      Visibility <- "10_DI_DATA_FS_332 FLW_OK"
      HorizontalMovement <- "82_To_HMI_FS332 Animation"
   Circle "Circle_69" at 573,764 size 8x8
      Visibility <- "10_DI_DATA_FS_332 FLW_OK"
      HorizontalMovement <- "82_To_HMI_FS332 Animation"
   Circle "Circle_70" at 712,763 size 8x8
      Visibility <- "10_DI_DATA_FS_332 FLW_OK"
      HorizontalMovement <- "82_To_HMI_FS332 Animation"
   Circle "Circle_74" at 822,763 size 8x8
      Visibility <- "10_DI_DATA_FS_332 FLW_OK"
      HorizontalMovement <- "82_To_HMI_FS332 Animation"
   Circle "Circle_75" at 828,691 size 8x8
      Visibility <- "10_DI_DATA_FS_332 FLW_OK"
      VerticalMovement <- "82_To_HMI_FS332 Animation"
   Circle "Circle_76" at 828,633 size 8x8
      Visibility <- "10_DI_DATA_FS_332 FLW_OK"
      VerticalMovement <- "82_To_HMI_FS332 Animation"
   Circle "Circle_77" at 763,613 size 8x8
      Visibility <- "10_DI_DATA_FS_332 FLW_OK"
      HorizontalMovement <- "82_To_HMI_FS332 Animation"
   Circle "Circle_78" at 845,515 size 10x10
      Visibility <- "10_DI_DATA_FS_332 FLW_OK"
      HorizontalMovement <- "82_To_HMI_FS332 Animation"
   Circle "Circle_79" at 856,642 size 10x10
      Visibility <- "10_DI_DATA_FS_332 FLW_OK"
      VerticalMovement <- "82_To_HMI_FS332 Animation"
   Circle "Circle_80" at 856,765 size 10x10
      Visibility <- "10_DI_DATA_FS_332 FLW_OK"
      VerticalMovement <- "82_To_HMI_FS332 Animation"
   Circle "Circle_55" at 179,684 size 7x7
      Visibility <- "10_DI_DATA_CV358_OPN"
      HorizontalMovement <- "82_To_HMI_P304 Animation"
   Circle "Circle_83" at 318,685 size 7x7
      Visibility <- "10_DI_DATA_CV358_OPN"
      DiagonalMovement <- "82_To_HMI_P304 Animation"
   Circle "Circle_81" at 416,684 size 7x7
      Visibility <- "10_DI_DATA_CV358_OPN"
      DiagonalMovement <- "82_To_HMI_P304 Animation"
   Circle "Circle_56" at 485,684 size 7x7
      Visibility <- "10_DI_DATA_CV358_OPN"
      DiagonalMovement <- "82_To_HMI_P304 Animation"
   Circle "Circle_85" at 496,641 size 7x7
      Visibility <- "10_DI_DATA_CV358_OPN"
      DiagonalMovement <- "82_To_HMI_P304 Animation"
   Circle "Circle_86" at 426,634 size 7x7
      Visibility <- "10_DI_DATA_CV358_OPN"
      DiagonalMovement <- "82_To_HMI_P304 Animation"
   TextField "Text field_50" at 969,420 size 254x154; Text 'Please Make Sure the Energy and Water Supply are Present and Sufficient'
      Visibility <- "Warn To Start GCU-Last"
   Button "Button_5" at 928,406 size 343x378; TextOff 'Text'
      Visibility <- "Warn To Start GCU-Last"
   TextField "Text field_21" at 919,606 size 359x94; Text 'Instalation Start Confirmation Required for Re-Ox Stage'
      Visibility <- "Warn To Start GCU-Last"
   Button "Button_6" at 1004,717 size 200x55; TextOff 'CONFIRM'; Authorization "Operate"
      on Press: function_b14e0dd5("80_From_HMI_GCU Start Confirmed", 0)
      Visibility <- "Warn To Start GCU-Last"
   TextField "Text field_51" at 914,433 size 366x124; Text 'Please Make Sure the Energy and Water Supply are Present and Sufficient'
      Visibility <- "Warn To Start GCU-Last"
   IOField "I/O field_37" at 1070,718 size 79x29; Authorization "Commissioning"; FormatPattern 999; Unit  step
      ProcessValue <- "2110_BTCS_CNTRL_DB_BTCS_STEP"
   Button "HmiScreenItemData_18" at 930,718 size 137x29; TextOn 'Back'; TextOff 'BWTS Step'
   Button "HmiScreenItemData_51" at 930,753 size 137x29; TextOn 'Back'; TextOff 'BWTS State'
   IOField "I/O field_38" at 1070,753 size 79x29; Authorization "Commissioning"; FormatPattern 9; Unit  state
      ProcessValue <- "2110_BTCS_CNTRL_DB_BTCS_STATE"
   TextField "Text field_64" at 497,462 size 54x22; Text '- OK -'
      Visibility <- "10_DI_DATA_LS_303_LO"
   GraphicView "Graphic view_76" at 53,433 size 168x182; Picture "Graphic_251"
   GraphicView "Graphic view_102" at 12,304 size 58x63; Picture "Graphic_162"
   GraphicView "Graphic view_13" at 724,163 size 182x22; Picture "Graphic_151"
   GraphicIOField "Graphic I/O field_3" at 188,659 size 60x65; PictureList "Pump Ani"
      ProcessValue <- "10_DI_DATA_P_304_ENBLD"
   GraphicView "Graphic view_18" at 240,683 size 253x11; Picture "Graphic_156"
   GraphicView "Graphic view_89" at 303,257 size 10x13; Picture "Graphic_147"
   GraphicView "Graphic view_59" at 962,301 size 302x22; Picture "Graphic_151"
   GraphicView "Graphic view_5" at 827,163 size 102x22; Picture "Graphic_151"
   GraphicView "Graphic view_69" at 124,683 size 68x11; Picture "Graphic_156"
   GraphicView "Graphic view_85" at 235,296 size 33x35; Picture "Graphic_178"
   GraphicView "Graphic view_1" at 259,128 size 301x502; Picture "Graphic_150"
   GraphicView "Graphic view_6" at 870,257 size 18x22; Picture "Graphic_154"
   GraphicView "Graphic view_9" at 689,257 size 188x11; Picture "Graphic_156"
   GraphicView "Graphic view_11" at 424,625 size 12x91; Picture "Graphic_152"
   GraphicView "Graphic view_10" at 424,628 size 19x28; Picture "Graphic_157"
   GraphicView "Graphic view_12" at 440,636 size 106x11; Picture "Graphic_156"
   GraphicView "Graphic view_14" at 817,752 size 20x21; Picture "Graphic_159"
   GraphicView "Graphic view_16" at 635,761 size 188x13; Picture "Graphic_151"
   GraphicIOField "Graphic I/O field_1" at 573,615 size 60x65; PictureList "Pump Ani"
      ProcessValue <- "10_DI_DATA_P_303_ENBLD"
   GraphicView "Graphic view_19" at 471,636 size 106x11; Picture "Graphic_156"
   TextField "Text field_16" at 90,573 size 90x22; Text 'PGC Running'
      Visibility <- "10_DI_DATA_E_400_RUN"
   GraphicView "Graphic view_21" at 486,674 size 17x18; Picture "Graphic_153"
   GraphicView "Graphic view_22" at 494,642 size 10x41; Picture "Graphic_152"
   GraphicView "Graphic view_23" at 490,637 size 17x15; Picture "Graphic_161"
   GraphicView "Graphic view_24" at 630,636 size 87x11; Picture "Graphic_156"
   GraphicView "Graphic view_33" at 668,469 size 24x18; Picture "Graphic_155"
   GraphicView "Graphic view_34" at 668,508 size 24x18; Picture "Graphic_166"
   GraphicView "Graphic view_35" at 679,517 size 62x11; Picture "Graphic_156"
   GraphicView "Graphic view_36" at 668,486 size 12x30; Picture "Graphic_152"
   GraphicView "Graphic view_37" at 687,468 size 62x11; Picture "Graphic_156"
   GraphicView "Graphic view_38" at 741,468 size 106x11; Picture "Graphic_156"
   GraphicView "Graphic view_39" at 487,257 size 103x11; Picture "Graphic_156"
   GraphicView "Graphic view_40" at 422,102 size 140x11; Picture "Graphic_156"
   GraphicView "Graphic view_41" at 302,103 size 24x18; Picture "Graphic_155"
   GraphicView "Graphic view_43" at 558,103 size 19x18; Picture "Graphic_154"
   GraphicView "Graphic view_44" at 302,118 size 12x75; Picture "Graphic_152"
   GraphicView "Graphic view_45" at 302,183 size 12x75; Picture "Graphic_152"
   GraphicView "Graphic view_46" at 871,460 size 17x18; Picture "Graphic_153"
   GraphicView "Graphic view_47" at 879,426 size 10x41; Picture "Graphic_152"
   GraphicView "Graphic view_48" at 771,468 size 106x11; Picture "Graphic_156"
   GraphicView "Graphic view_49" at 879,358 size 10x91; Picture "Graphic_152"
   GraphicView "Graphic view_51" at 879,272 size 10x91; Picture "Graphic_152"
   GraphicView "Graphic view_53" at 574,257 size 126x11; Picture "Graphic_156"
   GraphicView "Graphic view_57" at 319,102 size 140x11; Picture "Graphic_156"
   GraphicView "Graphic view_58" at 1062,188 size 19x119; Picture "Graphic_147"
   TextField "Text field_6" at 995,322 size 50x16; Text 'CV-407'
   GraphicView "Graphic view_61" at 561,250 size 23x16; Picture "Graphic_168"
   GraphicView "Graphic view_62" at 567,179 size 10x77; Picture "Graphic_152"
   TextField "Text field_8" at 1103,322 size 50x16; Text 'CV-411'
   TextField "Text field_13" at 1115,180 size 60x22; Text 'Opened'
      Visibility <- "10_DI_DATA_CV409_OPN"
   TextField "Text field_17" at 582,680 size 42x16; Text 'P-303'
   GraphicView "Graphic view_66" at 508,761 size 188x13; Picture "Graphic_151"
   GraphicView "Graphic view_67" at 375,761 size 188x13; Picture "Graphic_151"
   GraphicView "Graphic view_31" at 424,748 size 12x38; Picture "Graphic_152"
   GraphicView "Graphic view_68" at 118,761 size 285x13; Picture "Graphic_151"
   GraphicView "Graphic view_70" at 826,617 size 12x146; Picture "Graphic_147"
   GraphicView "Graphic view_71" at 818,611 size 19x21; Picture "Graphic_169"
   GraphicView "Graphic view_73" at 14,359 size 19x222; Picture "Graphic_147"
   GraphicView "Graphic view_75" at 696,479 size 76x194; Picture "Graphic_173"
   GraphicView "Graphic view_72" at 760,610 size 68x13; Picture "Graphic_151"
   GraphicView "Graphic view_32" at 847,514 size 19x20; Picture "Graphic_169"
   GraphicView "Graphic view_77" at 759,513 size 97x13; Picture "Graphic_151"
   GraphicView "Graphic view_28" at 855,527 size 12x146; Picture "Graphic_147"
   GraphicView "Graphic view_79" at 855,649 size 12x130; Picture "Graphic_147"
   TextField "Text field_24" at 610,79 size 50x16; Text 'CV-405'
   TextField "Text field_27" at 820,266 size 48x16; Text 'FS-350'
   GraphicView "Graphic view_15" at 834,232 size 20x26; Picture "Graphic_79"
   TextField "Text field_40" at 813,209 size 70x22; Text 'No Flow'
      Visibility <- "10_DI_DATA_FS_350_FLW_OK"
   TextField "Text field_41" at 813,209 size 70x22; Text '- Flow -'
      Visibility <- "10_DI_DATA_FS_350_FLW_OK"
   GraphicView "Graphic view_8" at 558,596 size 10x11; Picture "Graphic_159"
   GraphicView "Graphic view_17" at 563,440 size 5x162; Picture "Graphic_147"
   GraphicView "Graphic view_25" at 558,275 size 10x11; Picture "Graphic_169"
   GraphicView "Graphic view_27" at 563,280 size 5x177; Picture "Graphic_147"
   GraphicView "Graphic view_29" at 486,602 size 78x5; Picture "Graphic_151"
   GraphicView "Graphic view_80" at 488,275 size 76x5; Picture "Graphic_151"
   IOField "I/O field_2" at 524,401 size 82x35; FormatPattern 999.9; Unit  %
      ProcessValue <- "12_AI_Data_LIT_304_SCALED"
   TextField "Text field_29" at 669,184 size 56x16; Text 'PIT-416'
   GraphicView "Graphic view_81" at 687,140 size 20x26; Picture "Graphic_36"
   TextField "Text field_25" at 752,442 size 56x16; Text 'TIT-408'
   TextField "Text field_30" at 512,199 size 56x16; Text 'TIT-406'
   GraphicView "Graphic view_82" at 530,137 size 20x26; Picture "Graphic_36"
   TextField "Text field_26" at 824,348 size 56x16; Text 'PIT-353'
   GraphicView "Graphic view_84" at 15,559 size 33x36; Picture "Graphic_177"
   TextField "Text field_7" at 750,184 size 50x16; Text 'CV-406'
   Bar "Bar_1" at 377,282 size 109x327; Unit  %; MinimumValue 0; MaximumValue 100
      ProcessValue <- "12_AI_Data_LIT_304_SCALED"
   TextField "Text field_48" at 16,624 size 112x20; Text 'PG Compressor'
      Appearance <- "10_DI_DATA_E_400_NOK"
   TextField "Text field_34" at 615,534 size 79x34; Text 'Heat Exchanger'
   TextField "Text field_35" at 551,697 size 100x34; Text 'Recirculation Pump'
   TextField "Text field_36" at 402,782 size 61x18; Text 'To Bilge'
   TextField "Text field_37" at 814,782 size 100x18; Text 'To Overboard'
   TextField "Text field_38" at 571,440 size 55x16; Text 'LIT-304'
   TextField "Text field_39" at 269,693 size 56x16; Text 'PIT-358'
   GraphicView "Graphic view_90" at 287,658 size 20x26; Picture "Graphic_36"
   TextField "Text field_28" at 704,774 size 56x16; Text 'PIT-348'
   GraphicView "Graphic view_83" at 722,736 size 20x26; Picture "Graphic_36"
   TextField "Text field_31" at 778,623 size 48x16; Text 'FS-332'
   GraphicView "Graphic view_91" at 801,585 size 20x26; Picture "Graphic_79"
   TextField "Text field_32" at 779,562 size 70x22; Text 'No Flow'
      Visibility <- "10_DI_DATA_FS_332 FLW_OK"
   TextField "Text field_42" at 779,562 size 70x22; Text '- Flow -'
      Visibility <- "10_DI_DATA_FS_332 FLW_OK"
   TextField "Text field_43" at 197,724 size 42x16; Text 'P-304'
   TextField "Text field_44" at 169,740 size 106x20; Text 'Booster Pump'
   GraphicView "Graphic view_2" at 553,163 size 182x22; Picture "Graphic_151"
   GraphicView "Graphic view_7" at 251,453 size 24x21; Picture "Graphic_107"
   TextField "Text field_46" at 225,501 size 86x16; Text 'E-400-PT002'
   TextField "Text field_47" at 132,408 size 86x16; Text 'E-400-TT002'
   GraphicView "Graphic view_87" at 234,321 size 19x128; Picture "Graphic_147"
   GraphicView "Graphic view_86" at 220,442 size 33x36; Picture "Graphic_159"
   IOField "I/O field_10" at 683,53 size 57x22; FormatPattern 999
      ProcessValue <- "12_AI_Data_CV_405_SCALED"
   IOField "I/O field_11" at 226,482 size 68x18; FormatPattern 999.9; Unit  Bar
      ProcessValue <- "12_AI_Data_E_400_PT002_SCALED"
   IOField "I/O field_13" at 663,119 size 68x18; FormatPattern 99.99; Unit  Bar
      ProcessValue <- "12_AI_Data_PIT_416_SCALED"
   IOField "I/O field_14" at 787,330 size 68x18; FormatPattern 99.99; Unit  Bar
      ProcessValue <- "12_AI_Data_PIT_353_SCALED"
   IOField "I/O field_15" at 704,426 size 68x18; FormatPattern 99.99; Unit  °C
      ProcessValue <- "12_AI_Data_TIT_408_SCALED"
   IOField "I/O field_16" at 698,717 size 68x18; FormatPattern 99.99; Unit  Bar
      ProcessValue <- "12_AI_Data_PIT_348_SCALED"
   IOField "I/O field_7" at 263,638 size 68x18; FormatPattern 99.99; Unit  Bar
      ProcessValue <- "12_AI_Data_PIT_358_SCALED"
   TextField "Text field_57" at 1021,112 size 90x32; Text 'Vent To Atmosphere'
   TextField "Text field_58" at 608,3 size 150x18; Text 'Vent To Atmosphere'
   IOField "I/O field_1" at 143,392 size 68x18; FormatPattern 999.9; Unit  °C
      ProcessValue <- "12_AI_Data_E_400_TE002_SCALED"
   GraphicView "Graphic view_93" at 491,492 size 24x21; Picture "Graphic_107"
   TextField "Text field_63" at 515,491 size 48x16; Text 'LS-303'
   TextField "Text field_66" at 497,462 size 54x22; Text 'Low Low'
      Visibility <- "10_DI_DATA_LS_303_LO"
   TextField "Text field_90" at 497,462 size 54x22; Text '-LOW-'
      Visibility <- "10_DI_DATA_LS_303_LO"
   GraphicView "Graphic view_94" at 99,304 size 58x63; Picture "Graphic_162"
   TextField "Text field_70" at 125,264 size 60x22; Text 'Opened'
      Visibility <- "10_DI_DATA_CV441_OPN"
   TextField "Text field_71" at 126,288 size 50x16; Text 'CV-441'
   GraphicView "Graphic view_95" at 103,278 size 19x41; Picture "Graphic_147"
   TextField "Text field_72" at 93,222 size 65x32; Text 'Ambient Air Inlet'
   GraphicView "Graphic view_96" at 86,364 size 36x39; Picture "Graphic_159"
   GraphicView "Graphic view_97" at 28,382 size 70x22; Picture "Graphic_151"
   TextField "Text field_69" at 125,264 size 60x22; Text 'Closed'
      Visibility <- "10_DI_DATA_CV441_CLSD"
   TextField "Text field_12" at 1115,180 size 60x22; Text 'Closed'
      Visibility <- "10_DI_DATA_CV409_CLSD"
   GraphicView "Graphic view_98" at 0,278 size 33x35; Picture "Graphic_169"
   GraphicView "Graphic view_99" at 856,330 size 23x20; Picture "Graphic_255"
   GraphicView "Graphic view_100" at 728,443 size 20x26; Picture "Graphic_36"
   TextField "Text field_18" at 950,356 size 149x23; Text 'Hazardous Area'
   GraphicView "Graphic view_4" at 1204,277 size 20x26; Picture "Graphic_36"
   IOField "I/O field_3" at 1172,257 size 89x18; FormatPattern s99.99; Unit  Bar
      ProcessValue <- "20_TANKS_IP_DATA_RIO_06_FIRST_TANK_DECK_IG_PRESS"
   TextField "Text field_20" at 1186,322 size 56x16; Text 'PIT-415'
   GraphicView "Graphic view_50" at 100,253 size 26x26; Picture "Graphic_261"
   GraphicView "Graphic view_74" at 549,146 size 18x54; Picture "Graphic_281"
   GraphicView "Graphic view_78" at 256,278 size 17x59; Picture "Graphic_281"
   GraphicView "Graphic view_101" at 213,397 size 23x20; Picture "Graphic_255"
   TextField "Text field_56" at 1229,342 size 44x32; Text 'To BWTS'
   TextField "Text field_60" at 661,356 size 94x23; Text 'Safe Area'
   IOField "I/O field_4" at 683,37 size 57x22; FormatPattern 999
      ProcessValue <- "16_AQ_Data_CV405_CNTRL"
   TextField "Text field_106" at 752,38 size 59x18; Text 'OPENED'
   GraphicView "Graphic view_103" at 14,298 size 19x22; Picture "Graphic_147"
   TextField "Text field_73" at 34,288 size 50x16; Text 'CV-401'
   TextField "Text field_74" at 30,264 size 60x22; Text 'Opened'
      Visibility <- "10_DI_Data_CV401_OPN"
   TextField "Text field_75" at 30,264 size 60x22; Text 'Closed'
      Visibility <- "10_DI_Data_CV401_CLSD"
   Button "HmiScreenItemData_13" at 4,669 size 121x40; TextOn 'IGG Plant'; TextOff 'Fresh Water System'
      on Release: ActivateScreen("Fresh Water System", 0)
      Appearance <- "10 DI_DATA_P305_ENBLD"
   Button "HmiScreenItemData_11" at 3,745 size 122x41; TextOn 'IGG Plant'; TextOff 'Cooling System'
      on Release: ActivateScreen("Cooling System", 0)
   TextField "Text field_22" at 90,573 size 90x22; Text 'PGC Loaded'
      Visibility <- "10_DI_DATA_E_400_RUN"
   Button "HmiScreenItemData_12" at 46,424 size 177x198; TextOn 'IGG Plant'; TextOff 'Text'
      on Release: ActivateScreen("PGC System", 0)
   GraphicView "Graphic view_54" at 588,60 size 19x108; Picture "Graphic_147"
   GraphicView "Graphic view_55" at 586,28 size 95x54; Picture "Graphic_167"
   GraphicView "Graphic view_56" at 588,8 size 19x33; Picture "Graphic_147"
   IOField "I/O field_12" at 506,119 size 68x18; FormatPattern 99.99; Unit  °C
      ProcessValue <- "12_AI_Data_TIT_406_SCALED"
   GraphicView "Graphic view_42" at 567,116 size 10x51; Picture "Graphic_152"
   TextField "Text field_76" at 618,40 size 30x22; Text 'A'
      Visibility <- "19_AUTO_CMNDS_Data_CV405_PID_MDLTG"
   GraphicView "Logo" at 1,1 size 219x60; Picture "Logo of IGG HMI"
   Button "HmiScreenItemData_1" at 1,50 size 150x43; TextOn 'Back'; TextOff 'Main Index'
      on Release: ActivateScreen("02 Main Index", 0)
   GraphicView "Graphic view_92" at 925,164 size 33x36; Picture "Graphic_169"
   Button "HmiScreenItemData_2" at 1128,64 size 150x43; TextOn 'Back'; TextOff 'GCU Setup'
      on Release: ActivateScreen("Inert Gas Conditioning Setup", 0)
   DateTimeField "HmiScreenItemData_17" at 1175,0 size 105x30
   DateTimeField "HmiScreenItemData" at 1175,30 size 105x30
   GraphicView "Graphic view_106" at 939,194 size 19x100; Picture "Graphic_147"
   GraphicView "Graphic view_104" at 940,285 size 33x37; Picture "Graphic_177"
   Button "HmiScreenItemData_9" at 930,410 size 340x30; TextOn 'Back'; TextOff 'GCU CONTROL'
      Visibility <- "150_GCU_LCL_CNTRL_DB_LCL_CNTRL_ACTV"
   Line "Line_2" at 1246,550 size 0x80
      Visibility <- "150_GCU_LCL_CNTRL_DB_LCL_CNTRL_ACTV"
   Line "Line_3" at 1080,630 size 166x0
      Visibility <- "150_GCU_LCL_CNTRL_DB_LCL_CNTRL_ACTV"
   Button "HmiScreenItemData_4" at 930,610 size 150x40; TextOn 'Back'; TextOff 'Stop'
      on Press: function_b14e0dd5("150_GCU_LCL_CNTRL_DB_STOP", 0)
      Visibility <- "150_GCU_LCL_CNTRL_DB_LCL_CNTRL_ACTV"
   Line "Line_7" at 1080,530 size 145x0
      Visibility <- "150_GCU_LCL_CNTRL_DB_LCL_CNTRL_ACTV"
   Circle "Circle_20" at 1225,510 size 40x40
      Appearance <- "150_GCU_LCL_CNTRL_DB_RUN_WITH_AIR"
      Visibility <- "150_GCU_LCL_CNTRL_DB_LCL_CNTRL_ACTV"
   Button "HmiScreenItemData_3" at 930,510 size 150x40; TextOn 'Back'; TextOff 'Start With Air'
      on Press: function_b14e0dd5("150_GCU_LCL_CNTRL_DB_STRT_AIR", 0)
      Visibility <- "150_GCU_LCL_CNTRL_DB_LCL_CNTRL_ACTV"
   Button "HmiScreenItemData_5" at 930,450 size 340x40; TextOn 'Back'; TextOff 'Start'; TextList "GCU_LCL"
      ProcessValue <- "150_GCU_LCL_CNTRL_DB_LCL_CNTRL_ACTV"
      on Press: InvertBit("150_GCU_LCL_CNTRL_DB_LCL_CNTRL_ACTV")
      Visibility <- "150_GCU_LCL_CNTRL_DB_LCL_CNTRL_ACTV"
   Button "HmiScreenItemData_6" at 930,560 size 150x40; TextOn 'Back'; TextOff 'Start With IG'
      on Press: function_b14e0dd5("150_GCU_LCL_CNTRL_DB_STRT_IG", 0)
      Visibility <- "150_GCU_LCL_CNTRL_DB_LCL_CNTRL_ACTV"
   Line "Line_6" at 1080,580 size 145x0
      Visibility <- "150_GCU_LCL_CNTRL_DB_LCL_CNTRL_ACTV"
   Circle "Circle_1" at 1225,560 size 40x40
      Appearance <- "150_GCU_LCL_CNTRL_DB_RUN_WITH_IG"
      Visibility <- "150_GCU_LCL_CNTRL_DB_LCL_CNTRL_ACTV"
   Button "HmiScreenItemData_7" at 930,660 size 240x40; TextOn 'Back'; TextOff 'Start With Air'; TextList "GTT_OPS"
      on Press: InvertBit("150_GCU_LCL_CNTRL_DB_OPN_ACTV_GTT_VLVS")
      ProcessValue <- "150_GCU_LCL_CNTRL_DB_OPN_ACTV_GTT_VLVS"
      Visibility <- "150_GCU_LCL_CNTRL_DB_LCL_CNTRL_ACTV"
   Circle "Circle_2" at 1225,660 size 40x40
      Appearance <- "150_GCU_LCL_CNTRL_DB_OPN_ACTV_GTT_VLVS"
      Visibility <- "150_GCU_LCL_CNTRL_DB_LCL_CNTRL_ACTV"
   Line "Line_14" at 1170,680 size 55x0
      Visibility <- "150_GCU_LCL_CNTRL_DB_LCL_CNTRL_ACTV"
   Group "Group_4" at 187,631 size 60x25
   Group "Group_6" at 573,588 size 60x25
   IOField "I/O field_34" at 664,96 size 66x23; FormatPattern 99.9; Unit  Bar
      Appearance <- "19_AUTO_CMNDS_Data_PIT402_Target"
      ProcessValue <- "19_AUTO_CMNDS_Data_PIT416_CMND_Target"
   Group "Group_7" at 214,1 size 373x50
   GraphicView "Graphic view_105" at 1184,288 size 96x48; Picture "Graphic_235"
   Button "HmiScreenItemData_10" at 1178,277 size 102x71; TextOn 'Back'; TextOff 'Text'
      on Press: ActivateScreen("Balast Water Treatment Plant", 0)
   GraphicView "Graphic view_108" at 2,208 size 95x48; Picture "Left Arow"
   Button "HmiScreenItemData_14" at 1,195 size 106x107; TextOn 'Back'; TextOff 'Text'
      on Press: ActivateScreen("Inert Gas Generator Plant", 0)
   Button "HmiScreenItemData_15" at 1,133 size 158x52; TextOn 'INERT GAS TRANSFER'; TextOff 'Inert Gas Transfer'; TextList "IG Transfer"; Authorization "Operating Mode"
      on Release: ActivateScreen("IG Transfer Mode", 0)
      ProcessValue <- "80_From_HMI_BWT_BYPASS"
   GraphicView "Graphic view_88" at 434,257 size 55x11; Picture "Graphic_151"
   GraphicView "Graphic view_3" at 429,258 size 15x16; Picture "Graphic_178"
   Group "Group_5" at 396,264 size 74x42
   Group "Group_9" at 591,11 size 604x305
   Group "Group_10" at 389,152 size 96x105
   Group "Group_11" at 239,299 size 243x195
   Group "Group_8" at 384,257 size 504x388
   Group "Group_12" at 260,515 size 606x260
   Group "Group" at 746,80 size 58x108; Picture "Graphic_72"
   TextField "Text field_33" at 744,96 size 60x22; Text 'Closed'
      Visibility <- "10_DI_DATA_CV406_CLSD"
   TextField "Text field_14" at 744,96 size 60x22; Text 'Opened'
      Visibility <- "10_DI_DATA_CV406_OPN"
   Group "Group_2" at 991,218 size 58x108; Picture "Graphic_72"
   TextField "Text field_45" at 989,239 size 60x22; Text 'Closed'
      Visibility <- "10_DI_DATA_CV407_CLSD"
   TextField "Text field_11" at 989,239 size 60x22; Text 'Opened'
      Visibility <- "10_DI_DATA_CV407_OPN"
   Group "Group_3" at 1096,218 size 58x108; Picture "Graphic_72"
   TextField "Text field_9" at 1097,239 size 60x22; Text 'Closed'
      Visibility <- "10_DI_DATA_CV411_CLSD"
   TextField "Text field_10" at 1097,239 size 60x22; Text 'Opened'
      Visibility <- "10_DI_DATA_CV411_OPN"
   GraphicView "Graphic view_60" at 1058,159 size 58x63; Picture "Graphic_162"
   GraphicView "Graphic view_65" at 1062,151 size 19x23; Picture "Graphic_147"
   TextField "Text field_5" at 1082,212 size 50x16; Text 'CV-409'
   TextField "Text field_1" at 460,713 size 60x22; Text 'Closed'
      Visibility <- "10_DI_DATA_CV341_CLSD"
   TextField "Text field_2" at 460,713 size 60x22; Text 'Opened'
      Visibility <- "10_DI_DATA_CV341_OPN"
   GraphicView "Graphic view_30" at 421,704 size 39x47; Picture "Graphic_162"
   TextField "Text field_4" at 434,743 size 50x16; Text 'CV-341'
   GraphicView "Graphic view_26" at 424,662 size 12x54; Picture "Graphic_152"
   Group "Group_13" at 179,634 size 324x58
   TextField "Text field_3" at 356,693 size 50x16; Text 'CV-358'
   Group "Group_1" at 359,634 size 43x62; Picture "Graphic_72"
   TextField "Text field_15" at 350,634 size 60x22; Text 'Closed'
      Visibility <- "10_DI_DATA_CV358_CLSD"
   TextField "Text field_23" at 350,634 size 60x22; Text 'Opened'
      Visibility <- "10_DI_DATA_CV358_OPN"
   Button "Button_1" at 655,120 size 84x92; TextOff 'Text'
      on Press: function_efd93a16("PGC Setpoint Protection", 400, 200, -1, -1, 1)
   Button "Button_4" at 578,3 size 84x99; TextOff 'Text'
      on Press: function_efd93a16("CV 405 Grafics", 300, 100, -1, -1, 1)
   Button "HmiScreenItemData_16" at 236,593 size 83x29; TextOn 'Back'; TextOff 'Temp-Trends'
      on Click: function_efd93a16("PGC Temperature Trends", 200, 100, -1, -1, 1)
   GraphicView "Graphic view_107" at 563,347 size 57x58; Picture "Graphic_302"
      Visibility <- "10_DI_DATA_EPB_8S1"
   Group "Group_14" at 914,406 size 366x378

screen "GCU Target Setpoints" 1280x800, template "Template"
   on GenerateScreen: "TitleUpdater"()
   Button "HmiScreenItemData_1" at 1,1 size 150x43; TextOn 'Back'; TextOff 'Commissioning'
      on Release: ActivateScreen("Commissioning Main Page", 0)
   AlarmView "Alarm view_1" at 0,777 size 1280x23
   TextField "Text field_37" at 20,239 size 300x30; Text 'GCU Control PLC (Rack 3)'
   TextField "Text field_1" at 810,239 size 450x30; Text 'PROCESS STEP RELATED SETPOINTS & TARGETS'
   TextField "Text field_82" at 100,299 size 220x22; Text 'LIT304 GCU LEVEL'
   IOField "I/O field_22" at 350,299 size 70x22; FormatPattern 999; Unit  %
      ProcessValue <- "12_AI_Data_LIT_304_SCALED"
   IOField "I/O field_23" at 450,299 size 75x22; Authorization "Parameter Change"; FormatPattern 999
      ProcessValue <- "84_Setpoints_LIT304_InitialFill_LowLow"
   IOField "I/O field_24" at 550,299 size 75x22; Authorization "Parameter Change"; FormatPattern 999
      ProcessValue <- "84_Setpoints_LIT304_InitialFill_Low"
   IOField "I/O field_25" at 952,299 size 75x22; Authorization "Parameter Change"; FormatPattern 999
      ProcessValue <- "84_Setpoints_LIT304_InitialFill_High"
   IOField "I/O field_26" at 1052,299 size 75x22; Authorization "Parameter Change"; FormatPattern 999
      ProcessValue <- "84_Setpoints_LIT304_InitialFill_HighHigh"
   TextField "Text field_22" at 20,299 size 53x22; Text 'IW800'
   TextField "Text field_90" at 350,272 size 70x22; Text 'Reading'
   TextField "Text field_23" at 450,272 size 75x22; Text 'Low Low'
   TextField "Text field_26" at 550,272 size 75x22; Text 'Low'
   TextField "Text field_27" at 952,272 size 75x22; Text 'High'
   TextField "Text field_28" at 1052,272 size 75x22; Text 'High High'
   TextField "Text field_41" at 100,272 size 220x22; Text 'Description'
   TextField "Text field_43" at 20,272 size 53x22; Text 'AI'
   IOField "I/O field_27" at 750,299 size 75x22; Authorization "Parameter Change"; FormatPattern 999
      ProcessValue <- "84_Setpoints_LIT304_InitialFill_Target"
   TextField "Text field_29" at 750,272 size 75x22; Text 'Target'
   TextField "Text field_30" at 1152,299 size 100x22; Text 'INITIAL FILL'
   IOField "I/O field_28" at 450,339 size 75x22; Authorization "Parameter Change"; FormatPattern 999
      ProcessValue <- "84_Setpoints_LIT304_Refill_LowLow"
   IOField "I/O field_29" at 550,339 size 75x22; Authorization "Parameter Change"; FormatPattern 999
      ProcessValue <- "84_Setpoints_LIT304_Refill_Low"
   IOField "I/O field_30" at 952,339 size 75x22; Authorization "Parameter Change"; FormatPattern 999
      ProcessValue <- "84_Setpoints_LIT304_Refill_High"
   IOField "I/O field_40" at 1052,339 size 75x22; Authorization "Parameter Change"; FormatPattern 999
      ProcessValue <- "84_Setpoints_LIT304_Refill_HighHigh"
   IOField "I/O field_43" at 650,339 size 75x22; Authorization "Parameter Change"; FormatPattern 999
      ProcessValue <- "84_Setpoints_LIT304_Refill_Target_Low"
   TextField "Text field_31" at 1152,339 size 100x22; Text 'RE-FILL'
   IOField "I/O field_44" at 650,299 size 75x22; Authorization "Parameter Change"; FormatPattern 999
      ProcessValue <- "84_Setpoints_LIT304_InitialFill_Target_Low"
   TextField "Text field_32" at 645,272 size 83x22; Text 'Target Low'
   IOField "I/O field_45" at 750,339 size 75x22; Authorization "Parameter Change"; FormatPattern 999
      ProcessValue <- "84_Setpoints_LIT304_Refill_Target"
   TextField "Text field_2" at 100,379 size 220x22; Text 'PIT416 GAS TO DECK PRESS'
   IOField "I/O field_1" at 350,379 size 70x22; FormatPattern 9.9; Unit  Barg
      ProcessValue <- "12_AI_Data_PIT_416_SCALED"
   TextField "Text field_6" at 20,379 size 53x22; Text 'IW810'
   IOField "I/O field_4" at 750,379 size 75x22; Authorization "Parameter Change"; FormatPattern 9.9; Unit  Barg
      ProcessValue <- "84_Setpoints_PIT416_Target"
   TextField "Text field_7" at 100,419 size 220x22; Text 'PIT358 FCW INLET PRESS'
   IOField "I/O field_2" at 350,419 size 70x22; FormatPattern 9.9; Unit  Barg
      ProcessValue <- "12_AI_Data_PIT_358_SCALED"
   IOField "I/O field_3" at 450,419 size 75x22; Authorization "Parameter Change"; FormatPattern 9.9; Unit  Barg
      ProcessValue <- "84_Setpoints_PIT358_InitialFill_LowLow"
   IOField "I/O field_5" at 550,419 size 75x22; Authorization "Parameter Change"; FormatPattern 9.9; Unit  Barg
      ProcessValue <- "84_Setpoints_PIT358_InitialFill_Low"
   IOField "I/O field_6" at 952,419 size 75x22; Authorization "Parameter Change"; FormatPattern 99.9; Unit  Barg
      ProcessValue <- "84_Setpoints_PIT358_InitialFill_High"
   IOField "I/O field_7" at 1052,419 size 75x22; Authorization "Parameter Change"; FormatPattern 99.9; Unit  Barg
      ProcessValue <- "84_Setpoints_PIT358_InitialFill_HighHigh"
   TextField "Text field_8" at 20,419 size 53x22; Text 'IW812'
   TextField "Text field_9" at 1152,419 size 100x22; Text 'INITIAL FILL'
   IOField "I/O field_8" at 450,459 size 75x22; Authorization "Parameter Change"; FormatPattern 9.9; Unit  Barg
      ProcessValue <- "84_Setpoints_PIT358_Refill_LowLow"
   IOField "I/O field_9" at 550,459 size 75x22; Authorization "Parameter Change"; FormatPattern 9.9; Unit  Barg
      ProcessValue <- "84_Setpoints_PIT358_Refill_Low"
   IOField "I/O field_10" at 952,459 size 75x22; Authorization "Parameter Change"; FormatPattern 99.9; Unit  Barg
      ProcessValue <- "84_Setpoints_PIT358_Refill_High"
   IOField "I/O field_11" at 1052,459 size 75x22; Authorization "Parameter Change"; FormatPattern 99.9; Unit  Barg
      ProcessValue <- "84_Setpoints_PIT358_Refill_HighHigh"
   TextField "Text field_10" at 1152,459 size 100x22; Text 'RE-FILL'
   TextField "Text field_3" at 100,499 size 220x22; Text 'PIT353 RECIRC FCW PRESS'
   IOField "I/O field_12" at 350,499 size 70x22; FormatPattern 9.9; Unit  Barg
      ProcessValue <- "12_AI_Data_PIT_353_SCALED"
   IOField "I/O field_13" at 450,499 size 75x22; Authorization "Parameter Change"; FormatPattern 9.9; Unit  Barg
      ProcessValue <- "84_Setpoints_PIT353_InitialFill_LowLow"
   IOField "I/O field_14" at 550,499 size 75x22; Authorization "Parameter Change"; FormatPattern 9.9; Unit  Barg
      ProcessValue <- "84_Setpoints_PIT353_InitialFill_Low"
   IOField "I/O field_15" at 952,499 size 75x22; Authorization "Parameter Change"; FormatPattern 9.9; Unit  Barg
      ProcessValue <- "84_Setpoints_PIT353_InitialFill_High"
   IOField "I/O field_20" at 1052,499 size 75x22; Authorization "Parameter Change"; FormatPattern 9.9; Unit  Barg
      ProcessValue <- "84_Setpoints_PIT353_InitialFill_HighHigh"
   TextField "Text field_4" at 20,499 size 53x22; Text 'IW816'
   TextField "Text field_11" at 1152,499 size 100x22; Text 'INITIAL FILL'
   IOField "I/O field_21" at 450,539 size 75x22; Authorization "Parameter Change"; FormatPattern 9.9; Unit  Barg
      ProcessValue <- "84_Setpoints_PIT353_Refill_LowLow"
   IOField "I/O field_31" at 550,539 size 75x22; Authorization "Parameter Change"; FormatPattern 9.9; Unit  Barg
      ProcessValue <- "84_Setpoints_PIT353_Refill_Low"
   IOField "I/O field_32" at 952,539 size 75x22; Authorization "Parameter Change"; FormatPattern 9.9; Unit  Barg
      ProcessValue <- "84_Setpoints_PIT353_Refill_High"
   IOField "I/O field_33" at 1052,539 size 75x22; Authorization "Parameter Change"; FormatPattern 9.9; Unit  Barg
      ProcessValue <- "84_Setpoints_PIT353_Refill_HighHigh"
   TextField "Text field_12" at 1152,539 size 100x22; Text 'RE-FILL'
   TextField "Text field_5" at 836,272 size 107x22; Text 'Safe Target'
   IOField "I/O field_16" at 854,379 size 75x22; Authorization "Parameter Change"; FormatPattern 9.99; Unit  Barg
      ProcessValue <- "84_Setpoints_PIT416_Target_Safe"
   Group "Group" at 455,41 size 373x50
   Button "HmiScreenItemData_8" at 469,45 size 355x40; TextOn 'Back'; TextOff 'Text'
   TextField "Screen title" at 455,41 size 373x50; Text 'Screen title'

Template "Template" 1280x800
   Button "HmiScreenItemData_12" at 953,4 size 80x35; TextOn 'WARNING'; TextOff 'Warning'
      on Release: ActivateScreen("04 Alarm Log", 0)
      Visibility <- "62_Warning_Data_WRNG_PRSNT"
   Button "HmiScreenItemData_14" at 1040,4 size 80x35; TextOn 'ALARM'; TextOff 'Alarm'
      on Release: ActivateScreen("04 Alarm Log", 0)
      Visibility <- "60_Alarm_Data_ALRM_PRSNT"
   Button "HmiScreenItemData_20" at 866,4 size 80x35; TextOn 'Back'; TextOff 'Lockout'
      on Click: SetBit("80_From_HMI_Reset_Alarms")
      on Press: function_b14e0dd5("80_From_HMI_RST_LOCKOUT", 0)
      Appearance <- "82_To_HMI_E-STOP LATCHED"
   Button "HmiScreenItemData_24" at 770,3 size 64x35; TextOn 'MUTE'; TextOff 'Mute'
      on Press: function_b14e0dd5("80_From_HMI_SLNCE_BZR", 0)
      Appearance <- "80_From_HMI_SLNCE_BZR"
   GraphicView "Graphic view_24" at 836,3 size 29x41; Picture "Graphic_138"
      Visibility <- "Buzzer"
   Group "Group_11" at 300,4 size 240x30
   Button "HmiScreenItemData_26" at 547,4 size 216x31; TextOn 'Back'; TextOff 'Text'
   IOField "I/O field_9" at 636,8 size 40x23; FormatPattern 99; Unit h
      ProcessValue <- "103_Main_Burner_DB_Hours burn_CV"
   IOField "I/O field_16" at 677,8 size 40x23; FormatPattern 99; Unit m
      ProcessValue <- "103_Main_Burner_DB_Minutes burn_CV"
   IOField "I/O field_19" at 718,8 size 40x23; FormatPattern 99; Unit s
      ProcessValue <- "103_Main_Burner_DB_Seconds burn_CV"
   GraphicView "Graphic view_80" at 544,-4 size 59x52; Picture "Graphic_130"
      Visibility <- "103_Main_Burner_DB_DN_OK"
   IOField "I/O field_35" at 595,8 size 40x23; FormatPattern 99; Unit d
      ProcessValue <- "103_Main_Burner_DB_Days burn_CV"
   AlarmView "Alarm view_1" at 0,777 size 1280x23
   Circle "Circle_46" at 266,6 size 26x26
      Appearance <- "IGG PLC HEART BEAT"
      Visibility <- "TRUE"
   Circle "Circle_1" at 235,6 size 26x26
      Visibility <- "TRUE"
      Appearance <- "Setpoint Override_DB_Set Pressure"
   Button "Button_8" at 300,4 size 240x30; TextOn 'IGGS Shutting Down'; TextOff 'IGGS Shutting down'
      Visibility <- "100_IGG_AUTO_SEQ_DB_CRNT_STEP"
   Button "Button_2" at 300,4 size 240x30; TextOn 'IGGS Starting Up'; TextOff 'IGGS Starting Up'
      Visibility <- "100_IGG_AUTO_SEQ_DB_CRNT_STEP"

screen "Inert Gas Generator Setup" 1280x800, template "Template"
   Circle "Circle_2" at 221,236 size 29x29
      Appearance <- "82_To_HMI_CRNT_MODE_IGG"
   Button "HmiScreenItemData_1" at 1,1 size 150x43; TextOn 'Back'; TextOff 'Main Index'
      on Release: ActivateScreen("02 Main Index", 0)
   Button "HmiScreenItemData_8" at 44,70 size 230x29; TextOn 'Back'; TextOff 'IGGS Mode of Operation'
   Circle "Circle_1" at 221,177 size 29x29
      Appearance <- "82_To_HMI_CRNT_MODE_IGG"
   Button "HmiScreenItemData_4" at 50,167 size 150x51; TextOn 'Back'; TextOff 'Manual'; Authorization "Operating Mode"
      on Press: function_b14e0dd5("80_From_HMI_Request_Manual(1)", 0)
   Circle "Circle_9" at 221,116 size 29x29
      Appearance <- "82_To_HMI_CRNT_MODE_IGG"
   TextField "Text field_1" at 54,547 size 182x20; Text 'Cooling System Overrun'
   TextField "Text field_3" at 54,511 size 89x20; Text 'Description'
   TextField "Text field_5" at 54,671 size 274x20; Text 'IGG Combustion Chamber Post Purge'
   TextField "Text field_6" at 347,511 size 68x20; Text 'Setpoint'
   Button "HmiScreenItemData_6" at 44,467 size 401x29; TextOn 'Back'; TextOff 'IGGS Settings'
   IOField "I/O field_4" at 345,542 size 90x30; Authorization "Commissioning"; FormatPattern 999; Unit  s
      ProcessValue <- "80_From_HMI_Cooling System Overrun"
   IOField "I/O field_6" at 345,665 size 90x30; Authorization "Commissioning"; FormatPattern 999; Unit  s
      ProcessValue <- "80_From_HMI_Post Purge Time"
   TextField "Text field_4" at 54,712 size 294x20; Text 'Air / Inert Gas Pressure (Pre-Ignition)'
   IOField "I/O field_1" at 345,707 size 90x30; Authorization "Commissioning"; FormatPattern 999; Unit  mBar
      ProcessValue <- "84_Setpoints_PIT402_Pilot_Target"
   TextField "Text field_13" at 293,112 size 93x21; Text 'Description'
   IOField "I/O field_13" at 463,150 size 226x30; FormatPattern 9999999999999999999999999999999999999999
      ProcessValue <- "db_time_sync_time_system_READ"
   Button "HmiScreenItemData_26" at 284,70 size 421x29; TextOn 'Back'; TextOff 'Time Setting'
   Button "HmiScreenItemData_24" at 291,192 size 166x30; TextOn 'Back'; TextOff 'Set System Time'; Authorization "Parameter Change"
      on Activate: function_cbf290fd(0, 0)
   Button "HmiScreenItemData_16" at 894,69 size 187x29; TextOn 'Back'; TextOff 'IO'
   Button "HmiScreenItemData_2" at 719,69 size 163x29; TextOn 'Back'; TextOff 'Runtime'
   Button "HmiScreenItemData_10" at 725,107 size 150x51; TextOn 'Back'; TextOff 'Reset AUTO'; Authorization "User administration"
      on Press: function_b14e0dd5("80_From_HMI_RST_AUT_SEQ(1)", 0)
      Appearance <- "80_From_HMI_RST_AUT_SEQ(1)"
   DateTimeField "Date/time field_1" at 463,192 size 226x30; Authorization "Parameter Change"
   TextField "Text field_14" at 314,156 size 142x20; Text 'System Time (UTC)'
   Button "HmiScreenItemData_49" at 44,348 size 401x29; TextOn 'Back'; TextOff 'Inert Gas Transfer Mode'
   Circle "Circle_21" at 400,386 size 26x26
      Appearance <- "80_From_HMI_BWT_BYPASS"
   Button "HmiScreenItemData_50" at 67,384 size 304x33; TextOn 'Back'; TextOff 'Ballast Water Treatment'
      on Press: InvertBit("80_From_HMI_BWT_BYPASS(1)"); ResetBit("80_From_HMI_CRG_BLNK_MODE(1)")
      Appearance <- "80_From_HMI_BWT_BYPASS(1)"
      ObjectEnable <- "100_GCU_AUTO_SEQ_DB_CRNT_STEP"
   Circle "Circle_22" at 400,424 size 26x26
      Appearance <- "80_From_HMI_CRG_BLNK_MODE"
   Button "HmiScreenItemData_51" at 67,422 size 304x33; TextOn 'Back'; TextOff 'Cargo Blanketing'
      on Press: InvertBit("80_From_HMI_CRG_BLNK_MODE(1)"); ResetBit("80_From_HMI_BWT_BYPASS(1)")
      Appearance <- "80_From_HMI_CRG_BLNK_MODE(1)"
      ObjectEnable <- "100_GCU_AUTO_SEQ_DB_CRNT_STEP"
   Button "HmiScreenItemData_23" at 50,106 size 150x51; TextOn 'Back'; TextOff 'Full Automation'; Authorization "Operating Mode"
      on Press: function_b14e0dd5("80_From_HMI_Request_Auto(1)", 0)
   Button "HmiScreenItemData_3" at 1129,1 size 150x43; TextOn 'I&A Compressor Ok'; TextOff 'Back'
      on Release: function_efd93a16()
   IOField "I/O field_2" at 345,748 size 90x30; Authorization "Commissioning"; FormatPattern 999; Unit  mBar
      ProcessValue <- "84_Setpoints_PIT402_Main_Target"
   TextField "Text field_7" at 54,753 size 302x20; Text 'Air / Inert Gas Pressure (Post-Ignition)'
   Button "HmiScreenItemData_7" at 50,228 size 150x51; TextOn 'Back'; TextOff 'FAT Mode'; Authorization "User administration"
      on Press: InvertBit("80_From_HMI_FAT_Mode"); function_b14e0dd5("80_From_HMI_Request_Auto(1)", 0)
   Button "HmiScreenItemData_11" at 725,226 size 150x51; TextOn 'Back'; TextOff 'IGG Standalone'; Authorization "Operating Mode"
      on Press: InvertBit("80_From_HMI_IGG_STND_ALN")
      Appearance <- "80_From_HMI_IGG_STND_ALN"
   Button "HmiScreenItemData_12" at 910,107 size 150x35; TextOn 'Back'; TextOff 'P301 Present'; TextList "P301 Present"; Authorization "Operating Mode"
      on Press: InvertBit("80_From_HMI_P301_PRSNT(1)")
      Appearance <- "80_From_HMI_P301_PRSNT(1)"
      ProcessValue <- "80_From_HMI_P301_PRSNT(1)"
   Button "HmiScreenItemData_13" at 910,181 size 150x35; TextOn 'Back'; TextOff 'CV312 Present'; TextList "CV312 Present"; Authorization "User administration"
      on Press: InvertBit("80_From_HMI_CV312_PRSNT")
      Appearance <- "80_From_HMI_CV312_PRSNT"
      ProcessValue <- "80_From_HMI_CV312_PRSNT"
   Button "HmiScreenItemData_14" at 910,218 size 150x35; TextOn 'Back'; TextOff 'CV431 Present'; TextList "CV431 Present"; Authorization "Operating Mode"
      on Press: InvertBit("80_From_HMI_CV431_PRSNT")
      Appearance <- "80_From_HMI_CV431_PRSNT"
      ProcessValue <- "80_From_HMI_CV431_PRSNT"
   Button "HmiScreenItemData_15" at 910,255 size 150x35; TextOn 'Back'; TextOff 'CV432 Present'; TextList "CV432 Present"; Authorization "Operating Mode"
      on Press: InvertBit("80_From_HMI_CV432_PRSNT")
      Appearance <- "80_From_HMI_CV432_PRSNT"
      ProcessValue <- "80_From_HMI_CV432_PRSNT"
   Button "HmiScreenItemData_18" at 725,166 size 150x51; TextOn 'Back'; TextOff 'Silence Buzzer'; Authorization "User administration"
      on Press: function_b14e0dd5("80_From_HMI_SLNCE_BZR", 0)
      Appearance <- "80_From_HMI_SLNCE_BZR"
   IOField "I/O field_7" at 596,369 size 93x43; Authorization "Commissioning"; FormatPattern 999; Unit  step
      ProcessValue <- "100_IGG_AUTO_SEQ_DB_CRNT_STEP"
   IOField "I/O field_8" at 598,426 size 93x43; Authorization "Commissioning"; FormatPattern 999; Unit  step
      ProcessValue <- "100_BC_AUTO_SEQ_DB_CRNT_STEP"
   Button "HmiScreenItemData_9" at 485,376 size 102x29; TextOn 'Back'; TextOff 'IGG PLC'
   Button "HmiScreenItemData_17" at 485,433 size 102x29; TextOn 'Back'; TextOff 'BC PLC'
   Button "HmiScreenItemData_19" at 700,376 size 563x29; TextOn 'Back'; TextOff 'IGG STEP'; TextList "STEP LIST IGG"
      ProcessValue <- "100_IGG_AUTO_SEQ_DB_CRNT_STEP"
   Button "HmiScreenItemData_20" at 700,433 size 563x29; TextOn 'Back'; TextOff 'IGG STEP'; TextList "STEP LIST BC"
      ProcessValue <- "100_BC_AUTO_SEQ_DB_CRNT_STEP"
   AlarmView "Alarm view_1" at 0,777 size 1280x23
   IOField "I/O field_9" at 618,295 size 60x30; Authorization "Commissioning"; FormatPattern 99; Unit  s
      ProcessValue <- "80_From_HMI_Beacon frequency"
   IOField "I/O field_10" at 619,332 size 60x30; Authorization "Commissioning"; FormatPattern 99; Unit  min
      ProcessValue <- "80_From_HMI_Buzzer reset time"
   TextField "Text field_9" at 489,301 size 138x20; Text 'Beacon frequency'
   TextField "Text field_10" at 489,337 size 100x20; Text 'Buzzer reset'
   TextField "Text field_11" at 974,670 size 257x27; Text 'Proportionate Component PID'
   TextField "Text field_15" at 974,704 size 257x27; Text 'Integrative Component PID'
   TextField "Text field_16" at 974,737 size 257x27; Text 'Derivative Component PID'
   TextField "Text field_17" at 976,486 size 153x27; Text 'GAIN'
   TextField "Text field_18" at 974,515 size 153x27; Text 'Integration Time'
   TextField "Text field_19" at 974,549 size 153x27; Text 'Derivation Time'
   TextField "Text field_20" at 976,584 size 153x27; Text 'Maximum opening'
   Group "Group_15" at 1129,515 size 112x34; Authorization "User administration"; Picture "Graphic_284"; FormatPattern 99
   Group "Group_16" at 1129,550 size 112x34; Authorization "User administration"; Picture "Graphic_284"; FormatPattern 99
   Group "Group_3" at 1129,480 size 112x34; Authorization "User administration"; Picture "Graphic_284"; FormatPattern 99
   Switch "Switch_8" at 1222,670 size 32x29; CaptionText 'Switch'; TextOn 'ON'; TextOff 'OFF'; Authorization "User administration"; PictureOff "Design_5_PilotLight_Green_Off"; PictureOn "Design_5_PilotLight_Green_On"
      on Change: InvertBit("84_Setpoints_P_ON")
      ProcessValue <- "84_Setpoints_P_ON"
   Switch "Switch_9" at 1222,704 size 32x29; CaptionText 'Switch'; TextOn 'ON'; TextOff 'OFF'; Authorization "User administration"; PictureOff "Design_5_PilotLight_Green_Off"; PictureOn "Design_5_PilotLight_Green_On"
      on Change: InvertBit("84_Setpoints_I_ON")
      ProcessValue <- "84_Setpoints_I_ON"
   Switch "Switch_10" at 1222,735 size 32x29; CaptionText 'Switch'; TextOn 'ON'; TextOff 'OFF'; Authorization "User administration"; PictureOff "Design_5_PilotLight_Green_Off"; PictureOn "Design_5_PilotLight_Green_On"
      on Change: InvertBit("84_Setpoints_D_ON")
      ProcessValue <- "84_Setpoints_D_ON"
   Group "Group_1" at 1129,618 size 112x34; Authorization "User administration"; Picture "Graphic_284"; FormatPattern 99
   TextField "Text field_21" at 976,618 size 153x27; Text 'Minimum opening'
   Circle "Circle_29" at 707,748 size 20x20
      Appearance <- "Evolving Setpoint_DB_LevelBetter"
   TextField "Text field_22" at 736,744 size 199x27; Text 'O2 content geting Better'
   Gauge "Gauge_2" at 456,468 size 239x239; UnitText '%'; CaptionText 'O2 Content'
      Visibility <- "80_From_HMI_CRG_BLNK_MODE"
      ProcessValue <- "12_AI_Data_E600O2ContentIn"
      MaximumValue <- "84_Setpoints_E600_CB_HighHigh"
   Button "Button_25" at 582,743 size 95x31; TextOn 'grafic'; TextOff 'GRAFIC'; PictureOff "imageedit_175_8204096749"
      on Click: function_efd93a16("CV 203 Grafics", 200, 100, -1, -1, 1)
   Gauge "Gauge_3" at 456,468 size 239x239; UnitText '%'; CaptionText 'O2 Content'
      Visibility <- "80_From_HMI_BWT_BYPASS"
      ProcessValue <- "12_AI_Data_E600O2ContentIn"
      MaximumValue <- "84_Setpoints_E600_BWT_HighHigh"
   Group "Group_2" at 1129,584 size 112x34; Authorization "User administration"; Picture "Graphic_284"; FormatPattern 99
   Button "HmiScreenItemData_21" at 910,144 size 150x35; TextOn 'Back'; TextOff 'P305 Present'; TextList "P305 Present"; Authorization "Operating Mode"
      on Press: InvertBit("80_From_HMI_P305_PRSNT")
      Appearance <- "80_From_HMI_P305_PRSNT"
      ProcessValue <- "80_From_HMI_P305_PRSNT"
   TextField "Text field_2" at 54,589 size 192x20; Text 'BWT O2 Content Setpoint'
   IOField "I/O field_5" at 345,583 size 90x30; Authorization "Commissioning"; FormatPattern 99.99; Unit %
      ProcessValue <- "84_Setpoints_E600_BWT_Target"
   TextField "Text field_8" at 54,630 size 154x20; Text 'Cargo Blanketing O2'
   IOField "I/O field_3" at 345,624 size 90x30; Authorization "Commissioning"; FormatPattern 99.99; Unit %
      ProcessValue <- "84_Setpoints_E600_CB_Target"
   Gauge "Gauge_1" at 699,468 size 239x239; UnitText '%'; CaptionText 'CV 203'
      ProcessValue <- "16_AQ_Data_CV203_CNTRL"
   Button "Button_1" at 698,313 size 133x31; TextOn 'Reset Whitness'; TextOff 'Reset Whitness'; PictureOff "imageedit_175_8204096749"
      on Press: function_b14e0dd5("Tag_1", 0); function_b14e0dd5("Tag_2", 0); function_b14e0dd5("Tag_3", 0); function_b14e0dd5("Tag_4", 0); function_b14e0dd5("Tag_5", 0)
      Visibility <- "user_group"
   GraphicView "Graphic view_22" at 1129,515 size 112x34; Picture "Graphic_284"
   IOField "D5_I/O field_2" at 1144,523 size 62x18; Authorization "User administration"; FormatPattern 99999
      ProcessValue <- "84_Setpoints_Integration Time"
   TextField "D5_Text field_2" at 1204,523 size 23x18; Text 'ms / km/h'
   GraphicView "Graphic view_23" at 1129,550 size 112x34; Picture "Graphic_284"
   IOField "D5_I/O field_3" at 1144,558 size 62x18; FormatPattern 99999
      ProcessValue <- "84_Setpoints_Derive Time"
   TextField "D5_Text field_3" at 1204,558 size 23x18; Text 'ms / km/h'
   GraphicView "Graphic view_25" at 1129,480 size 112x34; Picture "Graphic_284"
   IOField "D5_I/O field_10" at 1144,488 size 62x18; Authorization "User administration"; FormatPattern 99.9999
      ProcessValue <- "84_Setpoints_Gain"
   TextField "D5_Text field_10" at 1204,488 size 23x18; Text 'km/h'
   GraphicView "Graphic view_1" at 1129,618 size 112x34; Picture "Graphic_284"
   IOField "D5_I/O field_1" at 1144,626 size 62x18; Authorization "User administration"; FormatPattern 999
      ProcessValue <- "84_Setpoints_Min Opening"
   TextField "D5_Text field_1" at 1204,626 size 23x18; Text '% / km/h'
   GraphicView "Graphic view_2" at 1129,584 size 112x34; Picture "Graphic_284"
   IOField "D5_I/O field_5" at 1144,592 size 62x18; Authorization "User administration"; FormatPattern 999
      ProcessValue <- "84_Setpoints_Max Opening"
   TextField "D5_Text field_5" at 1204,592 size 23x18; Text '% / km/h'

